// TIA Portal project "Robot_ur_lab" (V15.1)

(* hardware
DEVICE "S7-1200 station_1"  S7-1200 Station
   slot 0: "Rack_0"  S7-1200 Rack  Rack  V1.0
   slot 1: "PLC_1"  CPU 1215C DC/DC/DC  6ES7 215-1AG40-0XB0  V4.2
DEVICE "HMI_1"  KTP400 Basic PN
   slot 0: "HMI_1"  KTP400 Basic PN  6AV2 123-2DB03-0AX0  15.1.0.0
   slot 1: "HMI_RT_1"  KTP400 Basic PN  6AV2 123-2DB03-0AX0  15.1.0.0
   slot 5: "HMI_1.IE_CP_1"  PROFINET Interface  15.0.1.0
      slot 1: "PROFINET Interface_1"  PROFINET Interface
         slot 1: "Port_1"  Port
*)

// ===== PLC "PLC_1"  CPU 1215C DC/DC/DC =====

VAR_GLOBAL   // PLC tag table "Default tag table"
   "Detector" AT %Q0.7 : Bool;
   "B_Inicio" AT %I0.6 : Bool;
   "Reset" AT %M12.6 : Bool;
   "Lectura_blancos" AT %MW8 : Int;
   "Lectura_negros" AT %MW0 : Int;
   "Input_Blanco" AT %MW10 : Int;
   "Input_Negro" AT %MW6 : Int;
   "Cuenta_Blanco" AT %MW4 : Int;
   "Cuenta_Negro" AT %MW2 : Int;
   "V_Reset" AT %M12.0 : Bool;
   "In_sensor" AT %I1.0 : Bool;
   "Enviar_cuenta_N" AT %Q0.6 : Bool;
   "Enviar_cuenta_B" AT %Q0.5 : Bool;
   "Robot_mod" AT %Q0.4 : Bool;
   "V_Pausa" AT %M12.1 : Bool;
   "V_Inicio" AT %M12.2 : Bool;
   "Robot_pos" AT %I0.1 : Bool;
   "Cuenta_terminada_B" AT %M12.3 : Bool;
   "timer_cuenta_B" AT %M12.4 : Bool;
   "Cuenta_terminada_N" AT %M12.5 : Bool;
   "Activar_aire" AT %I0.0 : Bool;
   "Relevador_aire" AT %Q0.1 : Bool;
   "B_Reset" AT %I0.5 : Bool;
   "timer_cuenta_N" AT %M12.7 : Bool;
   "Fin_programa" AT %I0.2 : Bool;
   "Detect_toogle" AT %MW13 : Int;
   "Detect_act_B" AT %M15.0 : Bool;
   "Detect_act_N" AT %M15.1 : Bool;
END_VAR

// folder: System blocks/Program resources

DATA_BLOCK "IEC_Timer_0_DB"   // DB1
{ S7_Optimized_Access := 'TRUE' }
AUTHOR : Simatic
FAMILY : IEC
NAME : IEC_TMR
VERSION : 1.0
// stored: InstanceOfName IEC_TIMER
"IEC_TIMER"
BEGIN
END_DATA_BLOCK

DATA_BLOCK "IEC_Timer_0_DB_1"   // DB2
{ S7_Optimized_Access := 'TRUE' }
AUTHOR : Simatic
FAMILY : IEC
NAME : IEC_TMR
VERSION : 1.0
// stored: InstanceOfName IEC_TIMER
"IEC_TIMER"
BEGIN
END_DATA_BLOCK

DATA_BLOCK "IEC_Timer_0_DB_2"   // DB3
{ S7_Optimized_Access := 'TRUE' }
AUTHOR : Simatic
FAMILY : IEC
NAME : IEC_TMR
VERSION : 1.0
// stored: InstanceOfName IEC_TIMER
"IEC_TIMER"
BEGIN
END_DATA_BLOCK

DATA_BLOCK "IEC_Counter_0_DB"   // DB4
{ S7_Optimized_Access := 'TRUE' }
AUTHOR : Simatic
FAMILY : IEC
NAME : CNTR
VERSION : 1.0
// stored: InstanceOfName IEC_COUNTER
"IEC_COUNTER"
BEGIN
END_DATA_BLOCK

DATA_BLOCK "IEC_Counter_0_DB_1"   // DB5
{ S7_Optimized_Access := 'TRUE' }
AUTHOR : Simatic
FAMILY : IEC
NAME : CNTR
VERSION : 1.0
// stored: InstanceOfName IEC_COUNTER
"IEC_COUNTER"
BEGIN
END_DATA_BLOCK

DATA_BLOCK "IEC_Counter_0_DB_2"   // DB6
{ S7_Optimized_Access := 'TRUE' }
AUTHOR : Simatic
FAMILY : IEC
NAME : CNTR
VERSION : 1.0
// stored: InstanceOfName IEC_COUNTER
"IEC_COUNTER"
BEGIN
END_DATA_BLOCK

DATA_BLOCK "IEC_Timer_0_DB_3"   // DB7
{ S7_Optimized_Access := 'TRUE' }
AUTHOR : Simatic
FAMILY : IEC
NAME : IEC_TMR
VERSION : 1.0
// stored: InstanceOfName IEC_TIMER
"IEC_TIMER"
BEGIN
END_DATA_BLOCK

DATA_BLOCK "IEC_Timer_0_DB_4"   // DB8
{ S7_Optimized_Access := 'TRUE' }
AUTHOR : Simatic
FAMILY : IEC
NAME : IEC_TMR
VERSION : 1.0
// stored: InstanceOfName IEC_TIMER
"IEC_TIMER"
BEGIN
END_DATA_BLOCK

DATA_BLOCK "IEC_Counter_0_DB_3"   // DB9
{ S7_Optimized_Access := 'TRUE' }
AUTHOR : Simatic
FAMILY : IEC
NAME : CNTR
VERSION : 1.0
// stored: InstanceOfName IEC_COUNTER
"IEC_COUNTER"
BEGIN
END_DATA_BLOCK

// folder: (top level)

ORGANIZATION_BLOCK "Main"   // OB1, LAD, ProgramCycle
TITLE = "Main Program Sweep (Cycle)"
{ S7_Optimized_Access := 'TRUE' }
VERSION : 0.1
   VAR_INPUT
      Initial_Call : Bool;   // Initial call of this OB
      Remanence : Bool;   // =True, if remanent data are available
   END_VAR
   VAR_TEMP   // added for the SCL form of the ladder/FBD networks
      _w1 : Bool;
      _w2 : Bool;
   END_VAR
BEGIN

REGION Network 1: Detección B o N
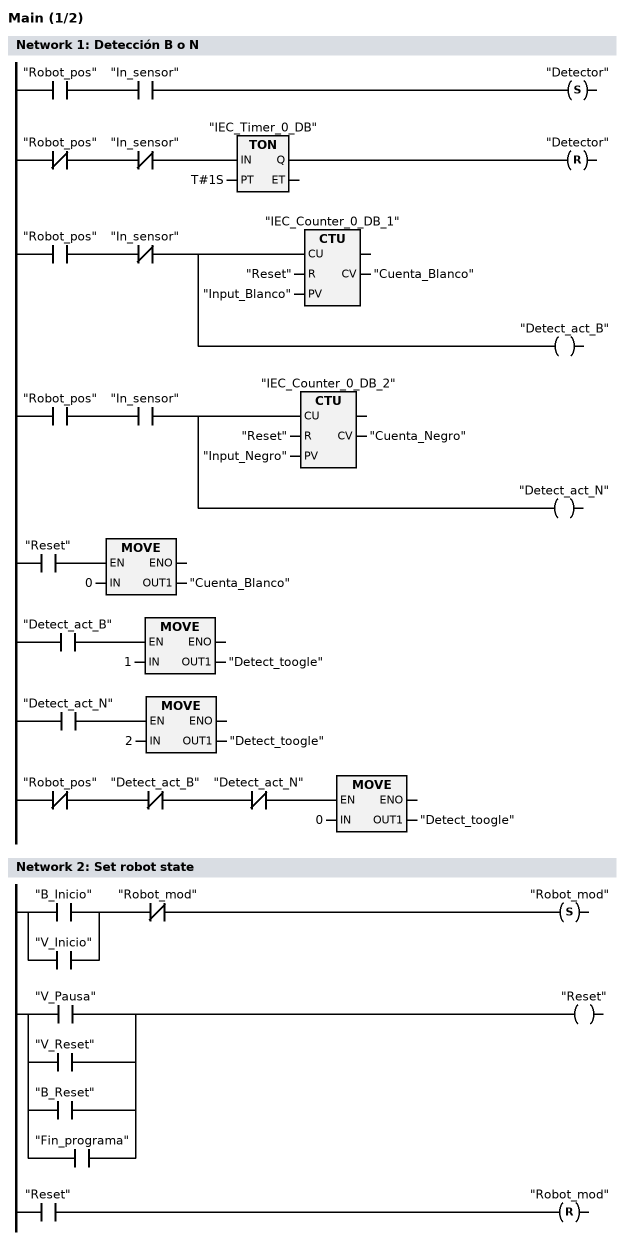
   IF "Robot_pos" AND "In_sensor" THEN "Detector" := TRUE; END_IF;
   "IEC_Timer_0_DB".TON(IN := NOT "Robot_pos" AND NOT "In_sensor", PT := T#1S);
   IF "IEC_Timer_0_DB".Q THEN "Detector" := FALSE; END_IF;
   #_w1 := "Robot_pos" AND NOT "In_sensor";
   "IEC_Counter_0_DB_1".CTU(CU := #_w1, R := "Reset", PV := "Input_Blanco", CV => "Cuenta_Blanco");
   "Detect_act_B" := #_w1;
   #_w2 := "Robot_pos" AND "In_sensor";
   "IEC_Counter_0_DB_2".CTU(CU := #_w2, R := "Reset", PV := "Input_Negro", CV => "Cuenta_Negro");
   "Detect_act_N" := #_w2;
   IF "Reset" THEN "Cuenta_Blanco" := 0; END_IF;
   IF "Detect_act_B" THEN "Detect_toogle" := 1; END_IF;
   IF "Detect_act_N" THEN "Detect_toogle" := 2; END_IF;
   IF NOT "Robot_pos" AND NOT "Detect_act_B" AND NOT "Detect_act_N" THEN "Detect_toogle" := 0; END_IF;
END_REGION

REGION Network 2: Set robot state
   RUNG wire#powerrail
      Contact( "B_Inicio" )
      wire#w1
      I_Contact( "Robot_mod" )
      S_Coil( "Robot_mod" )
   END_RUNG
   RUNG wire#powerrail
      Contact( "V_Inicio" )
   END_RUNG wire#w1
   RUNG wire#powerrail
      Contact( "V_Pausa" )
      wire#w2
      Coil( "Reset" )
   END_RUNG
   RUNG wire#powerrail
      Contact( "V_Reset" )
   END_RUNG wire#w2
   RUNG wire#powerrail
      Contact( "B_Reset" )
   END_RUNG wire#w2
   RUNG wire#powerrail
      Contact( "Fin_programa" )
   END_RUNG wire#w2
   RUNG wire#powerrail
      Contact( "Reset" )
      R_Coil( "Robot_mod" )
   END_RUNG
   // the same network as SCL:
   IF ("B_Inicio" OR "V_Inicio") AND NOT "Robot_mod" THEN "Robot_mod" := TRUE; END_IF;
   "Reset" := "V_Pausa" OR "V_Reset" OR "B_Reset" OR "Fin_programa";
   IF "Reset" THEN "Robot_mod" := FALSE; END_IF;
END_REGION

REGION Network 3: Enviar cuentas
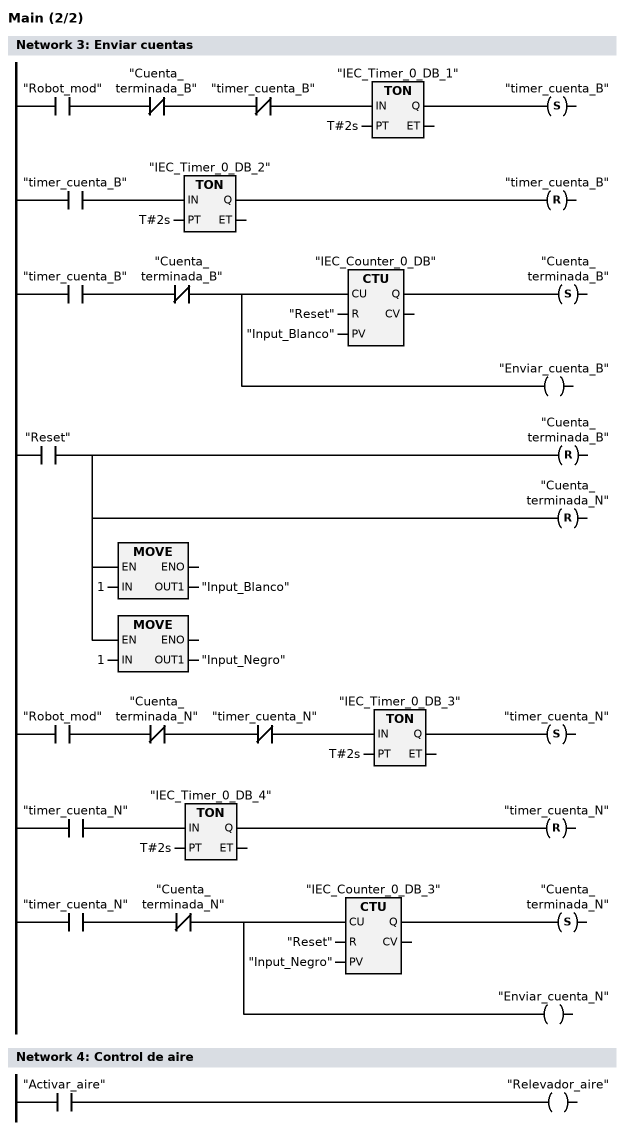
   "IEC_Timer_0_DB_1".TON(IN := "Robot_mod" AND NOT "Cuenta_terminada_B" AND NOT "timer_cuenta_B", PT := T#2s);
   IF "IEC_Timer_0_DB_1".Q THEN "timer_cuenta_B" := TRUE; END_IF;
   "IEC_Timer_0_DB_2".TON(IN := "timer_cuenta_B", PT := T#2s);
   IF "IEC_Timer_0_DB_2".Q THEN "timer_cuenta_B" := FALSE; END_IF;
   #_w1 := "timer_cuenta_B" AND NOT "Cuenta_terminada_B";
   "IEC_Counter_0_DB".CTU(CU := #_w1, R := "Reset", PV := "Input_Blanco");
   IF "IEC_Counter_0_DB".Q THEN "Cuenta_terminada_B" := TRUE; END_IF;
   "Enviar_cuenta_B" := #_w1;
   IF "Reset" THEN
       "Cuenta_terminada_B" := FALSE;
       "Cuenta_terminada_N" := FALSE;
       "Input_Blanco" := 1;
       "Input_Negro" := 1;
   END_IF;
   "IEC_Timer_0_DB_3".TON(IN := "Robot_mod" AND NOT "Cuenta_terminada_N" AND NOT "timer_cuenta_N", PT := T#2s);
   IF "IEC_Timer_0_DB_3".Q THEN "timer_cuenta_N" := TRUE; END_IF;
   "IEC_Timer_0_DB_4".TON(IN := "timer_cuenta_N", PT := T#2s);
   IF "IEC_Timer_0_DB_4".Q THEN "timer_cuenta_N" := FALSE; END_IF;
   #_w2 := "timer_cuenta_N" AND NOT "Cuenta_terminada_N";
   "IEC_Counter_0_DB_3".CTU(CU := #_w2, R := "Reset", PV := "Input_Negro");
   IF "IEC_Counter_0_DB_3".Q THEN "Cuenta_terminada_N" := TRUE; END_IF;
   "Enviar_cuenta_N" := #_w2;
END_REGION

REGION Network 4: Control de aire
   RUNG wire#powerrail
      Contact( "Activar_aire" )
      Coil( "Relevador_aire" )
   END_RUNG
   // the same network as SCL:
   "Relevador_aire" := "Activar_aire";
END_REGION
END_ORGANIZATION_BLOCK

(* ===== HMI "HMI_RT_1" =====
system functions are stored by id; their names below are inferred from use
connection "HMI_Connection_1": ETHERNET, SMART_S7_1200_OMS

HMI tags "Default tag table"
   "Tag_ScreenNumber" : UInt, internal
   "Detector_HMI" : Int = PLC Detect_toogle AT %MW13, 1 s
   "B_Inicio" : Bool = PLC V_Inicio AT %M12.2, 1 s
   "B_Pausa" : Bool = PLC V_Pausa AT %M12.1, 1 s
   "Input_Blanco" : Int = PLC Input_Blanco AT %MW10, 1 s
   "Input_Negro" : Int = PLC Input_Negro AT %MW6, 1 s
   "Cuenta_Blanco" : Int = PLC Cuenta_Blanco AT %MW4, 1 s
   "Cuenta_Negro" : Int = PLC Cuenta_Negro AT %MW2, 1 s
   "B_Reset" : Bool = PLC V_Reset AT %M12.0, 1 s

Template "Template_1" 480x272
   GraphicView "Logo" at 0,0 size 160x45; Picture "Logo of HMI_1"

screen "Color screen" 480x272, template "Template_1"
   TextField "Text field_1" at 202,93 size 70x27; Text 'Sensor'
   Rectangle "Rectangle_1" at 208,45 size 57x48
      Appearance <- "Detector_HMI"
   Button "Back" at 206,145 size 61x39; TextOn 'Back'; TextOff 'Inicio'
      on Press: SetTag("B_Inicio", 1)
      on Release: SetTag("B_Inicio", 0)
   Bar "Bar_1" at 30,110 size 80x120; MinimumValue 0; MaximumValue 8
      ProcessValue <- "Cuenta_Blanco"
   Bar "Bar_2" at 378,108 size 80x120; MinimumValue 0; MaximumValue 8
      ProcessValue <- "Cuenta_Negro"
   TextField "Text field_2" at 33,42 size 69x27; Text 'Blanco'
   TextField "Text field_4" at 378,42 size 63x27; Text 'Negro'
   Button "Back_3" at 206,198 size 61x39; TextOn 'Back'; TextOff 'Reinicio'
      on Release: SetTag("B_Reset", 0)
      on Press: SetTag("B_Reset", 1)
   IOField "I/O field_1" at 362,69 size 96x32; FormatPattern s99999
      ProcessValue <- "Input_Negro"
   IOField "I/O field_2" at 24,66 size 96x32; FormatPattern s99999
      ProcessValue <- "Input_Blanco"
*)